// Mitsubishi GX Works2 project: ZhaoQing_FenRong_Debug   PLC: Q06UDEH (continued)
           ELSE
   	        	H750Switch2io.xExitEnable:= H750Conveyor5IO.xEmpty;
    	        H750Conveyor5IO.xLoad:= H750Switch2ConveyorIn.xNextRun ;
            END_IF;
           	                                          
           H750ImportConveyor3IO.xLoad:=H750Switch2ConveyorOut.xNextRun AND m_iH750Switch2Select=1 ;
   	       H750ImportConveyor4IO.xLoad:=H750Switch2ConveyorOut.xNextRun AND m_iH750Switch2Select=2 ;
   	       IF  H750ImportConveyor3IO.xEmpty =0 AND H750ImportConveyor4IO.xEmpty =0 AND XCF AND XD0 THEN
   	       	H750ImportCylinder2IO.xMDIExe:=1;
   	       	H750ImportCylinder2IO.iDestinationPos:=2;
   	       	H750ImportConveyor3IO.xPutInto:=0;
   	       	H750ImportConveyor4IO.xPutInto:=0;
   	       END_IF;
   	       IF g_xImport2Force THEN (* 2巷道单框强制入库*)
   	       	H750ImportCylinder2IO.xMDIExe:=1;
   	       	H750ImportCylinder2IO.iDestinationPos:=2;
   	       	H750ImportConveyor3IO.xPutInto:=0;
   	       	H750ImportConveyor4IO.xPutInto:=0;   
   	       	END_IF;	       
   	       IF NOT XCF AND NOT XD0 THEN
   	       		H750ImportCylinder2IO.xMDIExe:=1;
   	       		H750ImportCylinder2IO.iDestinationPos:=1;
   	       END_IF;
   	       IF LDP(TRUE,H750ImportCylinder2IO.iCurrentPos=1 AND NOT H750ImportConveyor3IO.xCWPresent AND NOT H750ImportConveyor4IO.xCWPresent) THEN   	       	
   	       		H750ImportConveyor3IO.xPutInto:=1;
   	       		H750ImportConveyor4IO.xPutInto:=1;
   	       END_IF;        
      (*3巷道*)   
   			IF LDP(TRUE,H750Switch2ConveyorIn.xNextRun) THEN
  				H750Conveyor5IO.iProductCategory:= H750Switch2ConveyorIn.iProductCategory;  
  			END_IF;
         	H750Conveyor5IO.xUnload:=H750Conveyor6IO.xEmpty;
         	H750Conveyor6IO.xLoad:=H750Conveyor5IO.xNextRun;
   			IF LDP(TRUE,H750Conveyor5IO.xNextRun) THEN
  				H750Conveyor6IO.iProductCategory:= H750Conveyor5IO.iProductCategory;  
  			END_IF;             
            H750Switch3IO.xEntryEnable:=H750Conveyor6IO.xNextRun;
           (*分流信息传递到巷道3的顶升移载处*)
           H750Conveyor6IO.xUnload:=H750Switch3ConveyorIn.xEmpty;
           IF LDP(TRUE,H750Conveyor6IO.xNextRun) THEN
           	H750Switch3ConveyorIn.iProductCategory:=H750Conveyor6IO.iProductCategory;
           END_IF;
           (*分流信息显示为本巷道，启动顶升移载*)
           IF H750Switch3ConveyorIn.iProductCategory=4 THEN
           	H750Switch3IO.xSwithEnable:=1;
           ELSE
           	H750Switch3IO.xSwithEnable:=0;
           END_IF;
           (*双料入库，优先选择1 ，当1结束后恢复到0，2秒 ，然后再跳到2,0状态用来复位移载的出料*) 
          m_tonSwitch3NOSeleteDelay(IN:= m_iH750Switch3Select=0 ,PT:= t#2S ,Q:=m_xSwitch3NoSeleteDelay,ET:= m_tSwitch3NOSeleteDelayCurrentTi);
         IF   m_xSwitch3NoSeleteDelay THEN
         	m_xSwitch3SeleteDelay:=1;
         END_IF;
         IF ldf(TRUE, H750ImportConveyor5IO.xEmpty)  OR ldf(TRUE,H750ImportConveyor6IO.xEmpty) THEN
         	m_xSwitch3SeleteDelay:=0;
         END_IF;
   (*        m_tonSwitch1SeleteDelay(IN:= m_xSwitch1NOSeleteDelay  ,PT:= t#10S ,Q:= m_xSwitch1SeleteDelay ,ET:= m_tSwitch1SeleteDelayCurrentTime );     *)      
           IF H750ImportConveyor5IO.xEmpty AND  m_xSwitch3SeleteDelay   THEN
           		m_iH750Switch3Select:=1;
	           	ELSIF NOT H750ImportConveyor5IO.xEmpty AND H750ImportConveyor6IO.xEmpty AND m_xSwitch3SeleteDelay  THEN
           	  	m_iH750Switch3Select:=2;
          	 ELSE
           		m_iH750Switch3Select:=0;
           END_IF;
           IF H750Switch3IO.xSwithEnable THEN
         	  H750Switch3io.xExitEnable:=((H750ImportConveyor5IO.xEmpty AND m_iH750Switch3Select=1) 
                                                          OR   (H750ImportConveyor6IO.xEmpty AND m_iH750Switch3Select=2)) AND H750ImportCylinder3IO.iCurrentPos=1;
           ELSE
                   ;
                   (*报警，分流信息不正确*)
            END_IF;
           	                                          
           H750ImportConveyor5IO.xLoad:=H750Switch3ConveyorOut.xNextRun AND m_iH750Switch3Select=1 ;
   	       H750ImportConveyor6IO.xLoad:=H750Switch3ConveyorOut.xNextRun AND m_iH750Switch3Select=2 ;
   	       IF  H750ImportConveyor5IO.xEmpty =0 AND H750ImportConveyor6IO.xEmpty =0 AND XD6 AND XD7 THEN
   	       	H750ImportCylinder3IO.xMDIExe:=1;
   	       	H750ImportCylinder3IO.iDestinationPos:=2;
   	       	H750ImportConveyor5IO.xPutInto:=0;
   	       	H750ImportConveyor6IO.xPutInto:=0;
   	       END_IF;
   	       IF g_xImport3Force THEN (*3巷道单框强制入库*)
   	       	H750ImportCylinder3IO.xMDIExe:=1;
   	       	H750ImportCylinder3IO.iDestinationPos:=2;
   	       	H750ImportConveyor5IO.xPutInto:=0;
   	       	H750ImportConveyor6IO.xPutInto:=0;   
   	       	END_IF;	       
   	       IF NOT XD6 AND NOT XD7 THEN
   	       		H750ImportCylinder3IO.xMDIExe:=1;
   	       		H750ImportCylinder3IO.iDestinationPos:=1;
   	       END_IF;
   	       IF LDP(TRUE,H750ImportCylinder3IO.iCurrentPos=1 AND NOT H750ImportConveyor5IO.xCWPresent AND NOT H750ImportConveyor6IO.xCWPresent) THEN   	       	
   	       		H750ImportConveyor5IO.xPutInto:=1;
   	       		H750ImportConveyor6IO.xPutInto:=1;
   	       END_IF;            
         
         
         (*空框回流*)
         IF NOT M881 THEN  (*空框A回流*)
	         H2500EmptyASwitchIO.xEntryEnable:= NOT M881;
	         H2500EmptyASwitchIO.xLiftCylinderExtendInit:=0;
         ELSE
         	H2500EmptyASwitchIO.xEntryEnable:= 0;
         END_IF;
         H2500EmptyASwitchIO.xSwithEnable:=1;
    IF Lifter6IO.iCurrentPos=2 AND X3D THEN
    	IF NOT M881 THEN(*空框A回流的时候使用顶升移载退出命令*)
         H2500EmptyASwitchIO.xExitEnable:=COnveyor6IO.xEmpty;
    	END_IF;
    	IF M881 THEN(*空框B回流的时候使用顶升移载顶升移载下料输送线下料命令*)
         H2500EmptyASwitchConveyorOut.xUnload:=COnveyor6IO.xEmpty;
         END_IF;
    ELSE
    	H2500EmptyASwitchIO.xExitEnable:=0;
    	H2500EmptyASwitchConveyorOut.xUnload:=0;
    END_IF;
    (*空框B回流*)
    IF M881 THEN
    	H2500EmptyBSwitchIO.xEntryEnable:=M881;
    	H2500EmptyASwitchIO.xLiftCylinderExtendInit:=1;
    ELSE
    	H2500EmptyBSwitchIO.xEntryEnable:=0;
    END_IF;
     H2500EmptyBSwitchIO.xSwithEnable:=1;
     H2500EmptyBSwitchIO.xExitEnable:=H2500EmptyASwitchConveyorOut.xEmpty;
     H2500EmptyASwitchConveyorOut.xLoad:=H2500EmptyBSwitchConveyorOut.xNextRun;
    COnveyor6IO.xLoad:=H2500EmptyASwitchConveyorOut.xNextRun;
	IF COnveyor6IO.xEmpty THEN
		Lifter6IO.xMDIExe:=1;
		Lifter6Io.iDestinationPos:=2;
	END_IF;
	IF conveyor6IO.xEmpty=0 THEN
		Lifter6Io.xMDIExe:=1;
		Lifter6io.iDestinationPos:=1;
	END_IF;
	IF Lifter6IO.iCurrentPos=1 AND X3C AND H850RotorIO.iCurrentPos=1 AND X39 THEN
		COnveyor6IO.xUnload:=H850RotorConveyorIO.xEmpty;
	ELSE
		COnveyor6IO.xUnload:=0;
	END_IF;
	H850RotorConveyorIO.xLoad:=COnveyor6IO.xNextRun;
	(*临时使用人工投入空框程序，等空框回流线体能用之后解除下面的程序注释*)
(*	IF H850RotorConveyorIO.xEmpty THEN
		H850RotorIO.xMDIExe:=1;
		H850RotorIO.iDestinationPos:=1;
	END_IF;
	IF H850RotorConveyorIO.xEmpty=0 THEN
		H850RotorIO.xMDIExe:=1;
		H850RotorIO.iDestinationPos:=2;
	END_IF;*)
	(*====================================================*)
	H850RotorConveyorIO.xPutInto:=X139;
	IF H850RotorIO.iCurrentPos=2 AND X38 THEN
		H850RotorConveyorIO.xUnload:=H850Switch3ConveyorIn.xEmpty AND H850Switch3ConveyorOut.xEmpty;
	ELSE
		H850RotorConveyorIO.xUnload:=0;
	END_IF;
	H850Switch3IO.xEntryEnable:=H850RotorConveyorIO.xNextRun;
	H850Switch3IO.xSwithEnable:=1;
END_IF;
    (*报警程序*)
(*报警*)
M500:=D2315=1;(*分容库入库分流读码失败*)
M501:=D2320=1;(*常温库入库分流读码失败*)
g_xAlarm:=M500 
                     OR M501;
(*复位*)
IF g_xReset THEN
	g_xCommissioning:=0;
END_IF;
END_PROGRAM

PROGRAM Start
IF g_xReset THEN
	SM50:=1;
ELSE
	SM50:=0;
END_IF;
CASE g_iState OF
	0: 
		g_xManual:=1;
		g_xAuto:=0;	
		g_xStackLampAmber:=1;
		g_xStackLampGreen:=0;
		g_xRemoteAuto:=0;
	1:
		g_xManual:=0;
		g_xAuto:=1;
		g_xStackLampGreen:=1;
		g_xStackLampAmber:=0;
		g_xRemoteAuto:=0;
	2:	
        g_xRemoteAuto:=1;
        g_xStackLampGreen:=1;
        g_xStackLampAmber:=0;
        g_xAuto:=0;
		g_xManual:=0;
END_CASE;
IF g_xLocalAutoStart THEN  
	g_iState:=1;
END_IF;

IF g_xStop OR g_xEStop=0 THEN 
	g_iState:=0;
END_IF;
IF g_xRemoteAutoStart THEN
	g_iState:=2;
END_IF;
IF g_xAlarm AND SM412 THEN
	g_xStackLampRed:=1;
	g_xBuzzer:=1;
ELSE
	g_xStackLampRed:=0;
	g_xBuzzer:=0;	
END_IF;
END_PROGRAM

FUNCTION_BLOCK Conveyor
VAR
  tRundelay : TIME;  (* 离开延时 *)
END_VAR
VAR_IN_OUT
  ConveyorMotor : ConveyorIO;  (* 输送线输入输出 *)
END_VAR
VAR
  iStep : INT;  (* 上料步骤 *)
  m_tUnloadTimer : TIME;  (* 下料计时器 *)
  m_tonLeaveDelay : TON;  (* 离开延时定时器 *)
  m_xLeaveDelayOut : BOOL;  (* 离开延时 *)
  m_tLeaveCurrentTime : TIME;
END_VAR
VAR CONSTANT
  LOAD_UNLOAD_TIME : TIME := T#30s;  (* 延时报警常量 *)
END_VAR
VAR
  m_tonUnloadAlam : TON;  (* 下料报警定时器 *)
  m_tonLoadDelay : TON;  (* 离开延时定时器 *)
  m_xLoadDelayOut : BOOL;  (* 离开延时 *)
  m_tLoadCurrentTime : TIME;
  m_xInitial : BOOL;  (* 初始化 *)
  m_tLoadTimer : TIME;  (* 上料延时当前时间 *)
END_VAR
(*////////////////////////////////////////////////////////////////////////////////////////////////////////////
//传输线控制FB块，可控制单方向线体，双向旋转线体，支持双向上下料            
//线体初始化后为空的情况下输入xLoad信号即可进行上料动作，使用xLoadCCW信号可反方向上料
//增加了产品信息和产品种类的储存，当传输线为空和上料进行标志位为零的情况下清除产品信息和产品种类
//使用方式是在置位xLoad信号后，把产品信息和产品种类传入，等下料后自动清零
//线体不为空的情况下使用xUnload信号可进行下料动作，物料有无传感器的下降沿后出发计时器，延时断开传输线旋转
//单方向传输线体把xLoadCCW、xUnloadCCW设置为零，双向线体上料方向和下料反向的,方向固定的 把xUnloadCCW设置为1
//双方向线体双向都能上下料的要根据上料的方向来设置xLoadCCW,xUnloadCCW
//增加工作中信号xBusy当电机正转 显示为工作中
//增加上下料超时报警，xLoadAlarm，xUnloadAlarm，设定时间在LOAD_UNLOAD_TIME常量上，现在设置的为30秒
//增加xPutInto信号，用于直接投入的物料，检测开关感应到后，直接进入下料流程，上升沿有效
//离开延时改为变量 iLeaveDelay 默认为0 离开检测开关离输送线尾端比较远的线体需要根据情况设定100ms为单位
增加初始化标志位，增加进入延时时间，初始化为进入延时时间为0 ，离开延时时间为2S，通过外围接口可以更改
//修改信息  修改后请增加版本
//YAO      V1.0
///////////////////////////////////////////////////////////////////////////////////////////////////////////
********************************************************)
IF NOT m_xInitial THEN
	ConveyorMotor.tLoadDelay:=T#100ms;
	ConveyorMotor.xNegLimit:=1;
	ConveyorMotor.xPosLimit:=1;
	ConveyorMotor.xSizeDeficientDetect:=0;
END_IF;
m_xInitial:=1;
IF g_xAuto THEN
CASE iStep OF
	0:
	ConveyorMotor.xMotorCW:=0;
	ConveyorMotor.xMotorCCW:=0;
	ConveyorMotor.xNextRun:=0;
IF g_xEStop AND NOT ConveyorMotor.xLimitAlarrm AND NOT ConveyorMotor.xOverWidthAlarm  THEN
	IF  ConveyorMotor.xCWPresent OR ConveyorMotor.xCCWPresent  THEN
		iStep:=3;
		ConveyorMotor.xEmpty:=0;
		ELSE
		iStep:=1;
		ConveyorMotor.xEmpty:=1;
	END_IF;
END_IF;		
	1: 
	IF ConveyorMotor.xLoad    
		AND ConveyorMotor.xMotorCW=0   
		AND ConveyorMotor.xMotorCCW=0   
		AND ConveyorMotor.xEmpty THEN	
		iStep:=2;
	END_IF;
	2: 
	IF ConveyorMotor.xloadCCW THEN
		ConveyorMotor.xMotorCCW:=1; 
		ConveyorMotor.xMotorCW:=0;
	ELSE
	    ConveyorMotor.xMotorCW:=1;  
		ConveyorMotor.xMotorCCW:=0;
	END_IF;
		m_tonLoadDelay(IN:= (ConveyorMotor.xCWPresent AND NOT ConveyorMotor.xloadCCW) 
		                                        OR (ConveyorMotor.xCCWPresent AND ConveyorMotor.xloadCCW) ,
		                               PT:= ConveyorMotor.tLoadDelay ,
		                               Q:= m_xLoadDelayOut ,
		                               ET:= m_tLoadTimer );
	    IF (m_xLoadDelayOut AND NOT ConveyorMotor.xSizeDeficientDetect)   (*无尺寸检测时  只检测一个开关*)
	    	OR (m_xLoadDelayOut AND ConveyorMotor.xSizeDeficientDetect(*有尺寸检测时  要检测两个开关*)
	    	                                          AND ConveyorMotor.xCCWPresent 
	    	                                          AND ConveyorMotor.xCWPresent)      THEN 	 
		    iStep:=3;
			    ELSIF (m_xLoadDelayOut 
		                       AND ConveyorMotor.xSizeDeficientDetect(*尺寸不足报警*)
	    	                  AND (NOT ConveyorMotor.xCCWPresent OR NOT ConveyorMotor.xCWPresent))  
	    THEN
	    	    ConveyorMotor.xOverWidthAlarm:=1;
	    	   iStep:=0;               
	    END_IF;
	    
	3:
	ConveyorMotor.xMotorCW:=0;
	ConveyorMotor.xMotorCCW:=0;
	ConveyorMotor.xEmpty:=0;
	IF ConveyorMotor.xUnload AND NOT ConveyorMotor.xOverWidthAlarm THEN 
		iStep:=4;
	END_IF;
	4:	
	IF ConveyorMotor.xUnloadCCW THEN   
		ConveyorMotor.xMotorCCW:=1;  
		ConveyorMotor.xMotorCW:=0;
		ELSE
	    ConveyorMotor.xMotorCW:=1;  
		ConveyorMotor.xMotorCCW:=0;
	END_IF;
	ConveyorMotor.xNextRun:=1; 
	IF NOT ConveyorMotor.xUnload THEN 
		istep:=0;
	END_IF;
END_CASE;
IF LDP(TRUE,ConveyorMotor.xPutInto) THEN
	iStep:=0;
END_IF;
END_IF;
IF g_xManual THEN
	iStep:=0;

	IF ConveyorMotor.xForward 
		AND ConveyorMotor.xBackward=0 
		AND ConveyorMotor.xMotorCCW=0
		AND g_xEStop THEN
		ConveyorMotor.xMotorCW:=1;
		ConveyorMotor.xMotorCCW:=0;
		ELSE
		ConveyorMotor.xMotorCW:=0;
	END_IF;

	IF ConveyorMotor.xBackward 
		AND ConveyorMotor.xForward=0 
		AND ConveyorMotor.xMotorCW=0
		AND g_xEStop  THEN
		ConveyorMotor.xMotorCCW:=1;
		conveyormotor.xMotorCW:=0;
		ELSE
		ConveyorMotor.xMotorCCW:=0;
	END_IF;
END_IF;
IF ConveyorMotor.xMotorCCW        
	OR ConveyorMotor.xMotorCW THEN  
	ConveyorMotor.xBusy:=1;
	ELSE
	ConveyorMotor.xBusy:=0;
END_IF;
m_tonUnloadAlam(IN:= iStep=4,PT:= LOAD_UNLOAD_TIME,Q:= ConveyorMotor.xUnloadAlarm,ET:= m_tUnloadTimer );
(*//复位*)
IF (*g_xReset OR*)
	 (g_xResetSingle AND ConveyorMotor.iDeviceID=g_iDeviceIDSelect)THEN (*AND ConveyorMotor.iDeviceID=g_iDeviceIDSelect  THEN*)  (* //非正常情况下切断xNextRun不会复位，通过这个标志位会出发报警*)(*增加单体复位*)
	iStep:=0;
	ConveyorMotor.xNextRun:=0; 
	ConveyorMotor.xLimitAlarrm:=0;
	ConveyorMotor.xOverWidthAlarm:=0;
END_IF;
IF iStep=3 AND (NOT ConveyorMotor.xNegLimit OR NOT ConveyorMotor.xPosLimit) THEN
	ConveyorMotor.xOverWidthAlarm:=1;
END_IF;
IF ( ((ConveyorMotor.xloadCCW AND NOT ConveyorMotor.xNegLimit)            (*反转上料，碰到负限位*)
	OR  ( NOT ConveyorMotor.xloadCCW AND NOT ConveyorMotor.xPosLimit)) (*正转上料，碰到正限位*)
    AND iStep=2) (*上料过程*)
    OR
   ( iStep=4 (*下料过程*)
	AND( (ConveyorMotor.xUnloadCCW AND NOT ConveyorMotor.xPosLimit)  
	OR (NOT ConveyorMotor.xUnloadCCW AND NOT ConveyorMotor.xNegLimit)))    
    THEN
    ConveyorMotor.xLimitAlarrm:=1;
    iStep:=0;
END_IF;
END_FUNCTION_BLOCK

FUNCTION_BLOCK ShuttleCar
VAR_IN_OUT
  ShuttleCarInOut : ShuttleCarIO;
END_VAR
VAR
  m_tonBrakeDelay : TON;  (* 延时 *)
  m_tBrakeDelayCurrentTime : TIME;
  m_tonArriveDelay : TON;  (* 到达延时计时器 *)
  m_xInit : BOOL;  (* 初始化标志位 *)
  m_tonPauseDelay : TON;  (* 暂停减速 *)
  m_tPauseDelayCurrentTime : TIME;  (* 暂停延时当前时间 *)
  m_xArriveDelay : BOOL;  (* 到达延时 *)
  m_tArriveDelayCurrentTime : TIME;  (* 到达延时当前时间 *)
  m_tonOvertimeAlarm : TON;  (* 超时报警定时器 *)
  m_tOvertimeCurrentTime : TIME;  (* 超时报警当前时间 *)
END_VAR
(*******************************************************************
输送小车程序，可用于使用认址片控制位置的输送车程序，可用于控制提升机，
使用了限位捕捉程序防止小车惯性过大冲过限位后继续行走，捕捉程序采用反
转复位，这样设计有弊端可能反转复位后车的位置并没有回到限位以内,当两个
限位同时碰到的时候，会使运料小车进入死锁状态，通过xPassLimit来解开死锁，
可以在触摸屏中使用一个带权限的按钮来进行控制，配合ShuttleCarCurrentPos
函数来计算位置信息
增加自动开始后将当前位置置为零的信号防止设备停在两个位置开关的中间
修改信息  修改后请增加版本
2018-1-22增加到位延时：到位延时时间可以设置，适应双向到位的位置开关，通过调整延时时间让穿梭车停在到位开关的中间
增加气缸控制信号
增加抱闸延时
增加超时报警
YAO      V1.0
2018-1-22 YAO V1.1
********************************************************************)
IF NOT m_xInit THEN
	ShuttleCarInOut.tArriveDelay:=T#0s;   (*到位延时初始化为0*)
	ShuttleCarInOut.tBrakeDelay:=T#100ms;(*抱闸延时初始化为100ms*)
	ShuttleCarInOut.tSetOverTime:=T#60s;(*超时报警初始化为1分钟*)
	m_xInit:=1;
END_IF;
(*如果是气缸的话屏蔽限位和Ready信号*)
IF ShuttleCarInOut.xCylinder THEN
	ShuttleCarInOut.xPosLimit:=1;
	ShuttleCarInOut.xNegLimit:=1;
	ShuttleCarInOut.xReady:=1;
END_IF;
(*限位捕捉，防止冲过限位开关，反转后复位*)
ShuttleCarInOut.xPosLimitCatch:=LDF(TRUE,ShuttleCarInOut.xPosLimit) OR ShuttleCarInOut.xPosLimitCatch;
IF ShuttleCarInOut.xCCW THEN  
	ShuttleCarInOut.xPosLimitCatch:=0;
END_IF;

ShuttleCarInOut.xNegLimitCatch:=LDF(TRUE,ShuttleCarInOut.xNegLimit) OR ShuttleCarInOut.xNegLimitCatch;
(*松绳报警*)
IF LDP(TRUE,ShuttleCarInOut.xLooseDetect) THEN	
	ShuttleCarInOut.xLooseAlarm:=1;
END_IF;
(*提升复位报警*)
IF ShuttleCarInOut.xCW AND NOT  ShuttleCarInOut.xLooseDetect THEN   
	ShuttleCarInOut.xLooseAlarm:=0; 
END_IF;

IF ShuttleCarInOut.xCW THEN   
	ShuttleCarInOut.xNegLimitCatch:=0; 
END_IF;

IF ShuttleCarInOut.xPassLimit OR
	g_xReset OR   (*增加复位按钮*)
	(ShuttleCarInOut.xNegLimitCatch 
	AND ShuttleCarInOut.xPosLimitCatch)  THEN  
	ShuttleCarInOut.xNegLimitCatch:=0; 
	ShuttleCarInOut.xPosLimitCatch:=0;
	ShuttleCarInOut.xLooseAlarm:=0;
END_IF;
IF ShuttleCarInOut.xReady AND g_xEStop THEN
(*手动*)
    IF g_xManual THEN  
	    IF ShuttleCarInOut.xForward 
			AND ShuttleCarInOut.xBackward=0 
			AND ShuttleCarInOut.xCCW=0 
			AND ShuttleCarInOut.xPosLimitCatch=0  THEN
		    ShuttleCarInOut.xCW:=1;
		    ELSE
		    ShuttleCarInOut.xCW:=0;
	    END_IF;
	    IF ShuttleCarInOut.xBackward 
			AND ShuttleCarInOut.xForward=0 
			AND ShuttleCarInOut.xCW=0 
			AND ShuttleCarInOut.xNegLimitCatch=0 
			AND ShuttleCarInOut.xLooseAlarm=0
			AND G_xEStop THEN  
		    ShuttleCarInOut.xCCW:=1;
		    ELSE
		    ShuttleCarInOut.xCCW:=0;
	    END_IF;
    END_IF;
    (**********)
(*自动*)
  IF g_xAuto  THEN  
  	(*点动*)
 		IF LDP(TRUE,ShuttleCarInOut.xForward) THEN
 			ShuttleCarInOut.xMDIExe:=1;
			ShuttleCarInOut.iDestinationPos:=ShuttleCarInOut.iCurrentPos+1;
		END_IF;
		IF LDP(TRUE,ShuttleCarInOut.xBackward) THEN
			ShuttleCarInOut.xMDIExe:=1;
			ShuttleCarInOut.iDestinationPos:=ShuttleCarInOut.iCurrentPos-1;
		END_IF;	 
	(*>>>>>>>>>>>>>>>>>>>>>>>>>>>>>>>>>>>>>*)	
	  IF ShuttleCarInOut.xMDIExe AND ShuttleCarInOut.iDestinationPos<>0 THEN	
	    IF ShuttleCarInOut.iCurrentPos<ShuttleCarInOut.iDestinationPos AND ShuttleCarInOut.xPosLimitCatch=0 THEN   (*正转*)
			ShuttleCarInOut.xCW:=1;
			ShuttleCarInOut.xCCW:=0;
			ShuttleCarInOut.xMDIDone:=0;
		END_IF;

		IF ShuttleCarInOut.iCurrentPos>ShuttleCarInOut.iDestinationPos AND ShuttleCarInOut.xNegLimitCatch=0 AND ShuttleCarInOut.xLooseAlarm=0 THEN   (*反转*)
			ShuttleCarInOut.xCCW:=1;
			ShuttleCarInOut.xCW:=0;
			ShuttleCarInOut.xMDIDone:=0;
		END_IF;
	m_tonArriveDelay(IN:= ShuttleCarInOut.iCurrentPos=ShuttleCarInOut.iDestinationPos ,
	                                    PT:= ShuttleCarInOut.tArriveDelay ,
	                                    Q:= m_xArriveDelay ,
	                                    ET:= m_tArriveDelayCurrentTime);
	     (*到位延时时间可以设置，适应双向到位的位置开关，通过调整延时时间让穿梭车停在到位开关的中间*)
		IF m_xArriveDelay AND NOT ShuttleCarInOut.xCylinder THEN
			ShuttleCarInOut.xCW:=0;
			ShuttleCarInOut.xCCW:=0;
			ShuttleCarInOut.xMDIDone:=1;
			ELSE
			ShuttleCarInOut.xMDIDone:=0;
		END_IF;

		IF ShuttleCarInOut.xPosLimitCatch THEN
			ShuttleCarInOut.xCW:=0;
			ShuttleCarInOut.xMDIDone:=0;
		END_IF;

		IF ShuttleCarInOut.xNegLimitCatch THEN
			ShuttleCarInOut.xCCW:=0;
			ShuttleCarInOut.xMDIDone:=0;
		END_IF;
		ELSE
		ShuttleCarInOut.xCW:=0;
		ShuttleCarInOut.xCCW:=0;
		ShuttleCarInOut.xMDIDone:=0;
	  END_IF;
	END_IF;
	ELSE  (*无就绪信号   或急停的情况下*)
		ShuttleCarInOut.xCW:=0;
		ShuttleCarInOut.xCCW:=0;	
END_IF;
    (*抱闸延时*)
m_tonBrakeDelay(IN:= ShuttleCarInOut.xCW OR ShuttleCarInOut.xCCW,
                                    PT:= ShuttleCarInOut.tBrakeDelay,
                                    Q:=ShuttleCarInOut.xBrake ,
                                    ET:= m_tBrakeDelayCurrentTime);

(*自动上电后把当前位置清零，防止穿梭车不在开关位置*)
IF LDP(TRUE,g_xAuto) THEN
	ShuttleCarInOut.iCurrentPos:=0;
END_IF;
IF ShuttleCarInOut.xCW OR ShuttleCarInOut.xCCW THEN
	ShuttleCarInOut.xBusy:=1;
	ELSE
	ShuttleCarInout.xBusy:=0;
END_IF;

(*暂停，带延时减速斜坡，ShuttleCarInOut.xPauseRamp为减速斜坡输出位*)
m_tonPauseDelay(IN:=g_xPause,PT:= T#2s ,Q:=ShuttleCarInOut.xPauseRamp,ET:= m_tPauseDelayCurrentTime );
IF ShuttleCarInOut.xPauseRamp THEN
	ShuttleCarInOut.xCW:=0;
	ShuttleCarInOut.xCCW:=0;
	ShuttleCarInOut.xBrake:=0;
END_IF;
(*超时报警*)
m_tonOvertimeAlarm(IN:= ShuttleCarInOut.xMDIExe AND (ShuttleCarInOut.iCurrentPos<>ShuttleCarInOut.iDestinationPos) ,
                                           PT:= ShuttleCarInOut.tSetOverTime,
                                           Q:= ShuttleCarInOut.xOvertimeAlarm ,
                                           ET:= m_tOvertimeCurrentTime );
END_FUNCTION_BLOCK

FUNCTION ShuttleCarCurrentPosition
VAR_INPUT
  xPosition1 : BOOL;
  xPosition2 : BOOL;
  xPosition3 : BOOL;
END_VAR
(************************************
计算输送车当前位置的函数
**************************************)
IF xPosition1 THEN
	ShuttleCarCurrentPosition:=1;
END_IF;
IF xPosition2 THEN
	ShuttleCarCurrentPosition:=2;
END_IF;
IF xPosition3 THEN
	ShuttleCarCurrentPosition:=3;
END_IF;
END_FUNCTION

FUNCTION_BLOCK Switch
VAR_IN_OUT
  ConveyorEntryIO : ConveyorIO;
END_VAR
VAR
  ConveyorEntry : Conveyor;
  m_tonEntryBarDelay : TON;  (* 进入阻挡器延时 *)
  m_tEntryBarDelay : TIME;
  m_xEntryBarDelay : BOOL;
END_VAR
VAR_IN_OUT
  ConveyorExitIO : ConveyorIO;
END_VAR
VAR
  m_tonLiftCylinderDelay : TON;  (* 顶升延时 *)
  m_xLiftCylinderDelay : BOOL;
  m_tLiftCylinderDelay : TIME;
  m_tonExitBarDelay : TON;  (* 退出阻挡器延时 *)
  m_tExitBarDelay : TIME;
  m_xExitBarDelay : BOOL;
END_VAR
VAR_IN_OUT
  SwitchIO : SwitchIO;
END_VAR
VAR
  iStep : INT;
  ConveyorExit : Conveyor;
  m_xInitial : BOOL;
END_VAR
(**************************************************
顶升移载模块，抽象为一条输入输线 ，一条输出输送线
一个进入阻挡器，一个放出阻挡器，和一个顶升气缸的控制
程序思路比较混乱，接口不清晰，需要整改
直接放行的时候有问题
switchEnable =0的时候   离开线体的PutInto有问题
12-17日   V1.0
***************************************************)
ConveyorEntry(ConveyorMotor:=ConveyorEntryIO);
ConveyorExit(ConveyorMotor:=ConveyorExitIO);

IF NOT m_xInitial THEN
	
	m_xInitial:=1;
END_IF;
IF g_xAuto THEN
	CASE iStep OF
		0:(*初始化*)
		ConveyorEntryIO.xLoad:=0;
		ConveyorEntryIO.xUnload:=0;
		ConveyorEntryIO.xPutInto:=0;
		ConveyorExitIO.xLoad:=0;
		ConveyorExitIo.xUnload:=0;
		ConveyorExitIO.xPutInto:=0;
		SwitchIO.xEntryBarCylinderRetract:=0;
		SwitchIO.xExitBarCylinderRetract:=0;
		IF SwitchIO.xLiftCylinderExtendInit THEN
			SwitchIO.xLiftCylinderExtend:=1;
			SwitchIO.xLiftCylinderRetract:=0;
		    IF SwitchIO.xLiftCylinderExtendDetect THEN
			    iStep:=1;
		     END_IF; 
		ELSE
			SwitchIO.xLiftCylinderExtend:=0;
			SwitchIO.xLiftCylinderRetract:=1;	
		    IF SwitchIO.xLiftCylinderRetractDetect THEN
			    iStep:=1;
		    END_IF;		
		END_IF;
		1:(*上料*)
        IF SwitchIO.xEntryEnable AND ConveyorEntryIO.xEmpty AND ConveyorExitIO.xEmpty THEN
        	SwitchIO.xEntryBarCylinderRetract:=1;
        	ConveyorEntryIO.xLoad:=1;
        END_IF;
        IF ConveyorEntryIO.xEmpty=0 THEN
        	SwitchIO.xEntryBarCylinderRetract:=0;
        	ConveyorEntryIO.xLoad:=0;
        	ConveyorExitIO.xPutInto:=1;
        END_IF;
        IF m_xLiftCylinderDelay AND  SwitchIO.xSwithEnable THEN
        	 iStep:=2;
        END_IF;
        IF SwitchIO.xSwithEnable=0 AND m_xLiftCylinderDelay  THEN
        	 iStep:=3;
        END_IF;
		2:(*顶升*)
			SwitchIO.xExitBarCylinderRetract:=0;
		    IF SwitchIO.xLiftCylinderExtendInit THEN
			    SwitchIO.xLiftCylinderExtend:=0;
			    SwitchIO.xLiftCylinderRetract:=1;
		    ELSE
			    SwitchIO.xLiftCylinderExtend:=1;
			    SwitchIO.xLiftCylinderRetract:=0;			
		   END_IF;

		  IF SwitchIO.xLiftCylinderExtendInit THEN
		  	IF SwitchIO.xLiftCylinderRetractDetect THEN
		  		iStep:=4;
		  	END_IF;
		  	ELSE
		  	IF SwitchIO.xLiftCylinderExtendDetect THEN
		      iStep:=4; 
		  	END_IF;
		  END_IF;
		  3:(*放行*)	
		  	SwitchIO.xExitBarCylinderRetract:=1;
		  	ConveyorExitIO.xPutInto:=0;
		  	iStep:=4;
		  4:(*下料*)
		  (*通过出料传输线下料*)
		  IF SwitchIO.xExitEnable  AND m_xExitBarDelay AND NOT SwitchIO.xExitBarCylinderRetract  THEN		  
		  	ConveyorExitIO.xUnload:=1;
		  ELSE
		  	ConveyorExitIO.xUnload:=0;
		  END_IF;	
		   (*通过进料传输线下料*)
		  IF SwitchIO.xExitEnable  AND m_xExitBarDelay  AND SwitchIO.xExitBarCylinderRetract THEN		  
		  	ConveyorEntryIO.xUnload:=1;
		  ELSE
		  	ConveyorEntryIO.xUnload:=0;
		  END_IF;			    	
		  IF ConveyorExitIO.xEmpty OR ConveyorEntryIO.xEmpty  THEN
		  	ConveyorExitIO.xPutInto:=1;
		  	ConveyorEntryIO.xPutInto:=1;
			iStep:=0; 
		  END_IF;
	END_CASE;
        m_tonLiftCylinderDelay(IN:=NOT ConveyorEntryIO.xEmpty AND iStep=1 ,PT:= T#1S ,Q:= m_xLiftCylinderDelay ,ET:=m_tLiftCylinderDelay );
 		m_tonExitBarDelay(IN:=iStep=4 ,PT:= T#1s ,Q:= m_xExitBarDelay ,ET:= m_tExitBarDelay);
END_IF;
(*复位程序*)
IF (g_xResetSingle AND  (g_iDeviceIDSelect=ConveyorEntryIO.iDeviceID OR g_iDeviceIDSelect=ConveyorExitIO.iDeviceID))
	OR LDP(TRUE,SwitchIO.xLiftCylinderExtendInit) 
	OR LDF(TRUE,SwitchIO.xLiftCylinderExtendInit) 
	 THEN
	ConveyorEntryIO.xPutInto:=1;
	ConveyorExitIO.xPutInto:=1;
	iStep:=0;
END_IF;
IF g_xManual  THEN
	iStep:=0;
	ConveyorEntryIO.xLoad:=0;
    ConveyorEntryIO.xUnload:=0;
	ConveyorEntryIO.xPutInto:=0;
	ConveyorExitIO.xLoad:=0;
	ConveyorExitIo.xUnload:=0;
	ConveyorExitIO.xPutInto:=0;
	SwitchIO.xEntryBarCylinderRetract:=0;
	SwitchIO.xExitBarCylinderRetract:=0;
	IF SwitchIO.xEntryBarCylinderRetractButton THEN
		SwitchIO.xEntryBarCylinderRetract:=1;
	ELSE
		SwitchIO.xEntryBarCylinderRetract:=0;
	END_IF;
		IF SwitchIO.xExitBarCylinderRetractButton THEN
		SwitchIO.xExitBarCylinderRetract:=1;
	ELSE
		SwitchIO.xExitBarCylinderRetract:=0;
		END_IF;
		IF SwitchIO.xLiftCylinderExtendButton AND NOT SwitchIO.xLiftCylinderRetractButton THEN
			SwitchIO.xLiftCylinderExtend:=1;
			SwitchIO.xLiftCylinderRetract:=0;
		END_IF;
		IF NOT SwitchIO.xLiftCylinderExtendButton AND  SwitchIO.xLiftCylinderRetractButton THEN
			SwitchIO.xLiftCylinderExtend:=0;
			SwitchIO.xLiftCylinderRetract:=1;
		END_IF;		
	END_IF;
END_FUNCTION_BLOCK

FUNCTION_BLOCK ShuttleCarVelocityFB
VAR_INPUT
  xEnable : BOOL;  (* 使能 *)
  xMotorCW : BOOL;  (* 电机正转 *)
  xMotorCCW : BOOL;  (* 电机反转 *)
  xPosition1Switch : BOOL;  (* 位置1开关 *)
  xDecelerationSwitch : BOOL;  (* 减速开关 *)
  xPosition2Switch : BOOL;  (* 位置2开关 *)
END_VAR
VAR
  iFloor : INT;  (* 层数 *)
END_VAR
VAR_OUTPUT
  xHighSpeed : BOOL;
END_VAR
IF xEnable THEN
	(*电机旋转，并且在位置开关上的时候触发加速*)
	IF( LDP(TRUE,xMotorCW) AND xPosition1Switch ) OR (  LDP(TRUE,xMotorCCW) AND xPosition2Switch) THEN
		xHighSpeed:=1;
		iFloor:=0;
	END_IF;
	IF LDF(TRUE,xMotorCW) OR LDF(TRUE,xMotorCCW) THEN
		xHighSpeed:=0;
    END_IF;
	IF LDP(TRUE,xDecelerationSwitch) THEN
		iFloor:=iFloor+1;
	END_IF;
	IF iFloor=2 THEN
		xHighSpeed:=0;
		iFloor:=0;
	END_IF;
ELSE
    xHighSpeed:=0;
END_IF;
END_FUNCTION_BLOCK

FUNCTION_BLOCK BarCylinder
VAR_IN_OUT
  BarCylinderIO : BarCylinderIO;
END_VAR
VAR
  m_xInitial : BOOL;  (* 初始化 *)
  m_tonLoadDelay : TON;  (* 上料延时 *)
  m_xLoadDelay : BOOL;  (* 上料延时标志位 *)
  m_tLoadDelayCurrentTime : TIME;  (* 上料延时当前时间 *)
END_VAR
  (***********************************************************************
阻挡器模块，
由一个行程开关，一个阻挡器，一个倍速链输送电机组成
具有手动与自动模式
xEmpty显示当前为空料的状态
xUnload为卸料信号，连接下一设备的xEmpty信号
*************************************************************************)

IF NOT m_xInitial THEN
	BarCylinderIO.tLoadDelay:=T#5s;
	m_xInitial:=1;
END_IF;
IF g_xManual THEN    (*手动*)
	BarCylinderIO.xNextRun:=0;
	IF BarCylinderIO.xBarCylinderButton THEN
		BarCylinderIO.xBarCylinder:=1;
	ELSE
		BarCylinderIO.xBarCylinder:=0;
	END_IF;
	IF BarCylinderIO.xTransportMotorCWButton 
		AND NOT BarCylinderIO.xTransportMotorCCWButton 
		AND NOT BarCylinderIO.xTransportMotorCCW   THEN
		BarCylinderIO.xTransportMotorCW:=1;
	ELSE
		BarCylinderIO.xTransportMotorCW:=0;
	END_IF;
	IF BarCylinderIO.xTransportMotorCCWButton 
		AND NOT BarCylinderIO.xTransportMotorCWButton 
		AND NOT BarCylinderIO.xTransportMotorCW   THEN
		BarCylinderIO.xTransportMotorCCW:=1;
	ELSE
		BarCylinderIO.xTransportMotorCCW:=0;
	END_IF;
END_IF;
IF g_xAuto THEN(*自动*)
    IF BarCylinderIO.xUnload  AND NOT BarCylinderIO.xEmpty AND NOT BarCylinderIO.xNextRun THEN(*收到卸料命令，当阻挡器不为空时*)
    	BarCylinderIO.xBarCylinder:=1;
    	BarCylinderIO.xNextRun:=1;(*确保下料命令只执行一次，防止物料在输送过程中又有卸料命令导致多次卸料*)
    	BarCylinderIO.xTransportMotorCW:=1;
    END_IF;
    IF NOT  BarCylinderIO.xUnload  THEN
    	BarCylinderIO.xNextRun:=0;
    	BarCylinderIO.xBarCylinder:=0;
    END_IF;
    m_tonLoadDelay(IN:= BarCylinderIO.xPresentSwitch ,PT:= BarCylinderIO.tLoadDelay ,Q:= m_xLoadDelay,ET:= m_tLoadDelayCurrentTime );
    IF m_xLoadDelay OR  BarCylinderIO.xNextRun  THEN
    	BarCylinderIO.xEmpty:=0;
    ELSE
    	BarCylinderIO.xEmpty:=1;
    END_IF;
    (*如果为空，气缸顶起*)
   IF  BarCylinderIO.xEmpty  THEN
   	   BarCylinderIO.xBarCylinder:=0;
   END_IF;
   	IF BarCylinderIO.xLoad AND BarCylinderIO.xEmpty  THEN
		BarCylinderIO.xTransportMotorCW:=1;
   	END_IF;  
   	IF (BarCylinderIO.xLoad=0 OR BarCylinderIO.xEmpty=0)  AND (BarCylinderIO.xUnload=0 OR BarCylinderIO.xEmpty) THEN
   		BarCylinderIO.xTransportMotorCW:=0;
   	END_IF;
END_IF;  
IF BarCylinderIO.xEmpty AND BarCylinderIO.xLoad=0 THEN
	BarCylinderIO.iProductCategory:=0;
END_IF;

IF NOT g_xEStop THEN
	 BarCylinderIO.xTransportMotorCW:=0;
	 BarCylinderIO.xTransportMotorCCW:=0;
	 BarCylinderIO.xBarCylinder:=0;
END_IF;
END_FUNCTION_BLOCK

PROGRAM TCP
VAR
  m_ton6ReceiveHeartbeat : TON;
  m_t6RecHeartbeatCurrentTime : TIME;
  m_ton6ReceiveReConnect : TON;
  m_x6ReceiveReConnect : BOOL;
  m_t6ReceiveReConnectCurrentTime : TIME;
END_VAR
D220:=k18;
SP_SOCCINF( LDP(TRUE,SD1282.5) , "U0" , K6 , D140 ,D150);
SP_SOCSND( SM412 AND SD1282.5 , "U0" , K6 , D160, D220, M200 );
SP_SOCRCV( NOT M202  AND SD1282.5 , "U0" , K6, D310 , D420 ,M202);
D223.F:=SM413;
m_ton6ReceiveHeartbeat(IN:=NOT LDP(TRUE, D423.F) ,PT:= t#5S ,Q:= g_xQuarPackageRGVComFailed ,ET:= m_t6RecHeartbeatCurrentTime);
IF  g_xQuarPackageRGVComFailed THEN
	M202:=SM413;
	D420:=0;
	D421:=0;
	D422:=0;
	D423:=0;
	D424:=0;
END_IF;
END_PROGRAM

FUNCTION_BLOCK PiorityFb
VAR_INPUT
  xCondition1 : BOOL;  (* 条件1 *)
  xCondition2 : BOOL;  (* 条件2 *)
  xCondition3 : BOOL;  (* 条件3 *)
  xCondition4 : BOOL;  (* 条件4 *)
  xCondition5 : BOOL;  (* 条件5 *)
  xTaskComplete : BOOL;  (* 任务完成 *)
  xReset : BOOL;  (* 复位 *)
END_VAR
VAR
  xOccupy : BOOL;  (* 占用 *)
END_VAR
VAR_OUTPUT
  iPriority : INT;  (* 输出任务号 *)
END_VAR
VAR
  m_tonCondition1Delay : TON;
  m_xCondition1Delay : BOOL;
  m_tCondition1CurrentTime : TIME;
  arriTaskStack : ARRAY [0..5] OF INT;
  m_tonCondition2Delay : TON;
  m_xCondition2Delay : BOOL;
  m_tCondition2CurrentTime : TIME;
  m_tonCondition3Delay : TON;
  m_xCondition3Delay : BOOL;
  m_tCondition3CurrentTime : TIME;
  m_tonCondition4Delay : TON;
  m_xCondition4Delay : BOOL;
  m_tCondition4CurrentTime : TIME;
  m_tonCondition5Delay : TON;
  m_xCondition5Delay : BOOL;
  m_tCondition5CurrentTime : TIME;
  jj : INT;
END_VAR
(****************************************************************************)
(*
优先级功能块，存储5个条件的优先级，实现栈功能先入先出，
复位功能还有问题，
*)
(***************************************************************************)
m_tonCondition1Delay(IN:= xCondition1 AND NOT xReset ,PT:= T#1s,Q:= m_xCondition1Delay , ET:= m_tCondition1CurrentTime );
m_tonCondition2Delay(IN:= xCondition2 AND NOT xReset ,PT:= T#1s,Q:= m_xCondition2Delay , ET:= m_tCondition2CurrentTime );
m_tonCondition3Delay(IN:= xCondition3 AND NOT xReset ,PT:= T#1s,Q:= m_xCondition3Delay , ET:= m_tCondition3CurrentTime );
m_tonCondition4Delay(IN:= xCondition4 AND NOT xReset ,PT:= T#1s,Q:= m_xCondition4Delay , ET:= m_tCondition4CurrentTime );
m_tonCondition5Delay(IN:= xCondition5 AND NOT xReset ,PT:= T#1s,Q:= m_xCondition5Delay , ET:= m_tCondition5CurrentTime );

IF ldp(TRUE,m_xCondition1Delay) THEN
	FOR jj:=0 TO 5 BY 1 DO
		IF arriTaskStack[jj]=0 THEN
			arriTaskStack[jj]:=1;
			EXIT;
		END_IF;		
	END_FOR;
END_IF;

IF ldp(TRUE,m_xCondition2Delay) THEN
	FOR jj:=0 TO 5 BY 1 DO
		IF arriTaskStack[jj]=0 THEN
			arriTaskStack[jj]:=2;
			EXIT;
		END_IF;		
	END_FOR;
END_IF;

IF ldp(TRUE,m_xCondition3Delay) THEN
	FOR jj:=0 TO 5 BY 1 DO
		IF arriTaskStack[jj]=0 THEN
			arriTaskStack[jj]:=3;
			EXIT;
		END_IF;		
	END_FOR;
END_IF;

IF ldp(TRUE,m_xCondition4Delay) THEN
	FOR jj:=0 TO 5 BY 1 DO
		IF arriTaskStack[jj]=0 THEN
			arriTaskStack[jj]:=4;
			EXIT;
		END_IF;		
	END_FOR;
END_IF;

IF ldp(TRUE,m_xCondition5Delay) THEN
	FOR jj:=0 TO 5 BY 1 DO
		IF arriTaskStack[jj]=0 THEN
			arriTaskStack[jj]:=5;
			EXIT;
		END_IF;		
	END_FOR;
END_IF;

iPriority:=arriTaskStack[0];

IF 	LDP(TRUE, xTaskComplete) THEN
	FOR jj:=0 TO 4 BY 1 DO
		arriTaskStack[jj]:=arriTaskStack[jj+1];
	END_FOR;
		arriTaskStack[5]:=0;
END_IF;

IF LDP(TRUE,xReset) THEN
		FOR jj:=0 TO 5 BY 1 DO
		arriTaskStack[jj]:=0;
	END_FOR;
END_IF;
END_FUNCTION_BLOCK
